DATA_BLOCK "DB823_Error_Metering"   // DB823
TITLE = Faults general at plant and machine
{ S7_Optimized_Access := 'FALSE' }
VERSION : 0.1
   VAR
      FeedPump : Array[0..12] of "UDT1801_FLT_auxDrive";
      EdgeFilter : Array[0..12] of "UDT1801_EdgeFilter";
      MeteringPump : Array[0..12] of "UDT1853_FLT_MeteringPump";   // Metering pump
      Flow_Component : Array[0..12] of "UDT1822_FLT_PV_Flow";   // Process value flow component, mixing ratio
      Pressure_Component : Array[0..12] of "UDT1820_FLT_ProcessValue";   // Process value pressure at metering unit of component
      PrePressure_Component : Array[0..12] of "UDT1820_FLT_ProcessValue";   // Process value pressure at metering unit of component
      MicroMeteringUnit : Array[0..12] of "UDT1807_FaultMicroMeter";   // Micro metering unit ( Color)
      Temperature_HeatexchangerLP : Array[0..12] of "UDT1820_FLT_ProcessValue";   // Process value tempering heat exchanger
      Temperature_HeatexchangerHP : Array[0..12] of "UDT1820_FLT_ProcessValue";   // Process value tempering heat exchanger
      Temperature_Pump : Array[0..12] of "UDT1820_FLT_ProcessValue";   // Process value tempering pumps
      DifferencePressure : Array[0..12] of Struct
         BeforeEdge : "UDT1820_FLT_ProcessValue";
         BehindEdge : "UDT1820_FLT_ProcessValue";
         DifferenceEdge : "UDT1820_FLT_ProcessValue";
         BeforeHP : "UDT1820_FLT_ProcessValue";
         BehindHP : "UDT1820_FLT_ProcessValue";
         DifferenceHP : "UDT1820_FLT_ProcessValue";
      END_STRUCT;
      Heating : Array[0..12] of Struct
         Heating : Array[1..8] of "UDT1804_FLT_Controller";
      END_STRUCT;
   END_VAR
BEGIN
   FeedPump[0].FLT_Motorprotection := FALSE;
   FeedPump[0].FLT_FrequencyConverter := FALSE;
   FeedPump[0].FLT_MaxP_MaxLTripTray := FALSE;
   FeedPump[0].FLT_Dryrunsafety := FALSE;
   FeedPump[0].FLT_wrong_Timevalue := FALSE;
   FeedPump[0].FLT_MaxPressureDiff := FALSE;
   FeedPump[0].Mes_Min_temp := FALSE;
   FeedPump[0].FLT_MotorFan := FALSE;
   FeedPump[0].Mes_Min_Level := FALSE;
   FeedPump[0].FLT_No_Barrel := FALSE;
   FeedPump[0].Mes_No_Barrel := FALSE;
   FeedPump[0].Spare_1_3 := FALSE;
   FeedPump[0].Spare_1_4 := FALSE;
   FeedPump[0].Spare_1_5 := FALSE;
   FeedPump[0].Spare_1_6 := FALSE;
   FeedPump[0].Spare_1_7 := FALSE;
   FeedPump[1].FLT_Motorprotection := FALSE;
   FeedPump[1].FLT_FrequencyConverter := FALSE;
   FeedPump[1].FLT_MaxP_MaxLTripTray := FALSE;
   FeedPump[1].FLT_Dryrunsafety := FALSE;
   FeedPump[1].FLT_wrong_Timevalue := FALSE;
   FeedPump[1].FLT_MaxPressureDiff := FALSE;
   FeedPump[1].Mes_Min_temp := FALSE;
   FeedPump[1].FLT_MotorFan := FALSE;
   FeedPump[1].Mes_Min_Level := FALSE;
   FeedPump[1].FLT_No_Barrel := FALSE;
   FeedPump[1].Mes_No_Barrel := FALSE;
   FeedPump[1].Spare_1_3 := FALSE;
   FeedPump[1].Spare_1_4 := FALSE;
   FeedPump[1].Spare_1_5 := FALSE;
   FeedPump[1].Spare_1_6 := FALSE;
   FeedPump[1].Spare_1_7 := FALSE;
   FeedPump[2].FLT_Motorprotection := FALSE;
   FeedPump[2].FLT_FrequencyConverter := FALSE;
   FeedPump[2].FLT_MaxP_MaxLTripTray := FALSE;
   FeedPump[2].FLT_Dryrunsafety := FALSE;
   FeedPump[2].FLT_wrong_Timevalue := FALSE;
   FeedPump[2].FLT_MaxPressureDiff := FALSE;
   FeedPump[2].Mes_Min_temp := FALSE;
   FeedPump[2].FLT_MotorFan := FALSE;
   FeedPump[2].Mes_Min_Level := FALSE;
   FeedPump[2].FLT_No_Barrel := FALSE;
   FeedPump[2].Mes_No_Barrel := FALSE;
   FeedPump[2].Spare_1_3 := FALSE;
   FeedPump[2].Spare_1_4 := FALSE;
   FeedPump[2].Spare_1_5 := FALSE;
   FeedPump[2].Spare_1_6 := FALSE;
   FeedPump[2].Spare_1_7 := FALSE;
   FeedPump[3].FLT_Motorprotection := FALSE;
   FeedPump[3].FLT_FrequencyConverter := FALSE;
   FeedPump[3].FLT_MaxP_MaxLTripTray := FALSE;
   FeedPump[3].FLT_Dryrunsafety := FALSE;
   FeedPump[3].FLT_wrong_Timevalue := FALSE;
   FeedPump[3].FLT_MaxPressureDiff := FALSE;
   FeedPump[3].Mes_Min_temp := FALSE;
   FeedPump[3].FLT_MotorFan := FALSE;
   FeedPump[3].Mes_Min_Level := FALSE;
   FeedPump[3].FLT_No_Barrel := FALSE;
   FeedPump[3].Mes_No_Barrel := FALSE;
   FeedPump[3].Spare_1_3 := FALSE;
   FeedPump[3].Spare_1_4 := FALSE;
   FeedPump[3].Spare_1_5 := FALSE;
   FeedPump[3].Spare_1_6 := FALSE;
   FeedPump[3].Spare_1_7 := FALSE;
   FeedPump[4].FLT_Motorprotection := FALSE;
   FeedPump[4].FLT_FrequencyConverter := FALSE;
   FeedPump[4].FLT_MaxP_MaxLTripTray := FALSE;
   FeedPump[4].FLT_Dryrunsafety := FALSE;
   FeedPump[4].FLT_wrong_Timevalue := FALSE;
   FeedPump[4].FLT_MaxPressureDiff := FALSE;
   FeedPump[4].Mes_Min_temp := FALSE;
   FeedPump[4].FLT_MotorFan := FALSE;
   FeedPump[4].Mes_Min_Level := FALSE;
   FeedPump[4].FLT_No_Barrel := FALSE;
   FeedPump[4].Mes_No_Barrel := FALSE;
   FeedPump[4].Spare_1_3 := FALSE;
   FeedPump[4].Spare_1_4 := FALSE;
   FeedPump[4].Spare_1_5 := FALSE;
   FeedPump[4].Spare_1_6 := FALSE;
   FeedPump[4].Spare_1_7 := FALSE;
   FeedPump[5].FLT_Motorprotection := FALSE;
   FeedPump[5].FLT_FrequencyConverter := FALSE;
   FeedPump[5].FLT_MaxP_MaxLTripTray := FALSE;
   FeedPump[5].FLT_Dryrunsafety := FALSE;
   FeedPump[5].FLT_wrong_Timevalue := FALSE;
   FeedPump[5].FLT_MaxPressureDiff := FALSE;
   FeedPump[5].Mes_Min_temp := FALSE;
   FeedPump[5].FLT_MotorFan := FALSE;
   FeedPump[5].Mes_Min_Level := FALSE;
   FeedPump[5].FLT_No_Barrel := FALSE;
   FeedPump[5].Mes_No_Barrel := FALSE;
   FeedPump[5].Spare_1_3 := FALSE;
   FeedPump[5].Spare_1_4 := FALSE;
   FeedPump[5].Spare_1_5 := FALSE;
   FeedPump[5].Spare_1_6 := FALSE;
   FeedPump[5].Spare_1_7 := FALSE;
   FeedPump[6].FLT_Motorprotection := FALSE;
   FeedPump[6].FLT_FrequencyConverter := FALSE;
   FeedPump[6].FLT_MaxP_MaxLTripTray := FALSE;
   FeedPump[6].FLT_Dryrunsafety := FALSE;
   FeedPump[6].FLT_wrong_Timevalue := FALSE;
   FeedPump[6].FLT_MaxPressureDiff := FALSE;
   FeedPump[6].Mes_Min_temp := FALSE;
   FeedPump[6].FLT_MotorFan := FALSE;
   FeedPump[6].Mes_Min_Level := FALSE;
   FeedPump[6].FLT_No_Barrel := FALSE;
   FeedPump[6].Mes_No_Barrel := FALSE;
   FeedPump[6].Spare_1_3 := FALSE;
   FeedPump[6].Spare_1_4 := FALSE;
   FeedPump[6].Spare_1_5 := FALSE;
   FeedPump[6].Spare_1_6 := FALSE;
   FeedPump[6].Spare_1_7 := FALSE;
   FeedPump[7].FLT_Motorprotection := FALSE;
   FeedPump[7].FLT_FrequencyConverter := FALSE;
   FeedPump[7].FLT_MaxP_MaxLTripTray := FALSE;
   FeedPump[7].FLT_Dryrunsafety := FALSE;
   FeedPump[7].FLT_wrong_Timevalue := FALSE;
   FeedPump[7].FLT_MaxPressureDiff := FALSE;
   FeedPump[7].Mes_Min_temp := FALSE;
   FeedPump[7].FLT_MotorFan := FALSE;
   FeedPump[7].Mes_Min_Level := FALSE;
   FeedPump[7].FLT_No_Barrel := FALSE;
   FeedPump[7].Mes_No_Barrel := FALSE;
   FeedPump[7].Spare_1_3 := FALSE;
   FeedPump[7].Spare_1_4 := FALSE;
   FeedPump[7].Spare_1_5 := FALSE;
   FeedPump[7].Spare_1_6 := FALSE;
   FeedPump[7].Spare_1_7 := FALSE;
   FeedPump[8].FLT_Motorprotection := FALSE;
   FeedPump[8].FLT_FrequencyConverter := FALSE;
   FeedPump[8].FLT_MaxP_MaxLTripTray := FALSE;
   FeedPump[8].FLT_Dryrunsafety := FALSE;
   FeedPump[8].FLT_wrong_Timevalue := FALSE;
   FeedPump[8].FLT_MaxPressureDiff := FALSE;
   FeedPump[8].Mes_Min_temp := FALSE;
   FeedPump[8].FLT_MotorFan := FALSE;
   FeedPump[8].Mes_Min_Level := FALSE;
   FeedPump[8].FLT_No_Barrel := FALSE;
   FeedPump[8].Mes_No_Barrel := FALSE;
   FeedPump[8].Spare_1_3 := FALSE;
   FeedPump[8].Spare_1_4 := FALSE;
   FeedPump[8].Spare_1_5 := FALSE;
   FeedPump[8].Spare_1_6 := FALSE;
   FeedPump[8].Spare_1_7 := FALSE;
   FeedPump[9].FLT_Motorprotection := FALSE;
   FeedPump[9].FLT_FrequencyConverter := FALSE;
   FeedPump[9].FLT_MaxP_MaxLTripTray := FALSE;
   FeedPump[9].FLT_Dryrunsafety := FALSE;
   FeedPump[9].FLT_wrong_Timevalue := FALSE;
   FeedPump[9].FLT_MaxPressureDiff := FALSE;
   FeedPump[9].Mes_Min_temp := FALSE;
   FeedPump[9].FLT_MotorFan := FALSE;
   FeedPump[9].Mes_Min_Level := FALSE;
   FeedPump[9].FLT_No_Barrel := FALSE;
   FeedPump[9].Mes_No_Barrel := FALSE;
   FeedPump[9].Spare_1_3 := FALSE;
   FeedPump[9].Spare_1_4 := FALSE;
   FeedPump[9].Spare_1_5 := FALSE;
   FeedPump[9].Spare_1_6 := FALSE;
   FeedPump[9].Spare_1_7 := FALSE;
   FeedPump[10].FLT_Motorprotection := FALSE;
   FeedPump[10].FLT_FrequencyConverter := FALSE;
   FeedPump[10].FLT_MaxP_MaxLTripTray := FALSE;
   FeedPump[10].FLT_Dryrunsafety := FALSE;
   FeedPump[10].FLT_wrong_Timevalue := FALSE;
   FeedPump[10].FLT_MaxPressureDiff := FALSE;
   FeedPump[10].Mes_Min_temp := FALSE;
   FeedPump[10].FLT_MotorFan := FALSE;
   FeedPump[10].Mes_Min_Level := FALSE;
   FeedPump[10].FLT_No_Barrel := FALSE;
   FeedPump[10].Mes_No_Barrel := FALSE;
   FeedPump[10].Spare_1_3 := FALSE;
   FeedPump[10].Spare_1_4 := FALSE;
   FeedPump[10].Spare_1_5 := FALSE;
   FeedPump[10].Spare_1_6 := FALSE;
   FeedPump[10].Spare_1_7 := FALSE;
   FeedPump[11].FLT_Motorprotection := FALSE;
   FeedPump[11].FLT_FrequencyConverter := FALSE;
   FeedPump[11].FLT_MaxP_MaxLTripTray := FALSE;
   FeedPump[11].FLT_Dryrunsafety := FALSE;
   FeedPump[11].FLT_wrong_Timevalue := FALSE;
   FeedPump[11].FLT_MaxPressureDiff := FALSE;
   FeedPump[11].Mes_Min_temp := FALSE;
   FeedPump[11].FLT_MotorFan := FALSE;
   FeedPump[11].Mes_Min_Level := FALSE;
   FeedPump[11].FLT_No_Barrel := FALSE;
   FeedPump[11].Mes_No_Barrel := FALSE;
   FeedPump[11].Spare_1_3 := FALSE;
   FeedPump[11].Spare_1_4 := FALSE;
   FeedPump[11].Spare_1_5 := FALSE;
   FeedPump[11].Spare_1_6 := FALSE;
   FeedPump[11].Spare_1_7 := FALSE;
   FeedPump[12].FLT_Motorprotection := FALSE;
   FeedPump[12].FLT_FrequencyConverter := FALSE;
   FeedPump[12].FLT_MaxP_MaxLTripTray := FALSE;
   FeedPump[12].FLT_Dryrunsafety := FALSE;
   FeedPump[12].FLT_wrong_Timevalue := FALSE;
   FeedPump[12].FLT_MaxPressureDiff := FALSE;
   FeedPump[12].Mes_Min_temp := FALSE;
   FeedPump[12].FLT_MotorFan := FALSE;
   // 3232 more start values not shown
END_DATA_BLOCK

DATA_BLOCK "DB824_Error_MH_CP"   // DB824
TITLE = Faults mixinghead and cleaning piston
{ S7_Optimized_Access := 'FALSE' }
VERSION : 0.1
   VAR
      MH_Control : Array[0..16] of "UDT1842_FLT_MH_Control";
      CPiston : Array[0..16] of "UDT1871_FLT_CPiston";
      Temperature : Array[1..6, 0..16] of "UDT1820_FLT_ProcessValue";
      Pressure : Array[1..6, 0..16] of "UDT1820_FLT_ProcessValue";
      SteeringPiston : Array[0..16] of "UDT1820_FLT_ProcessValue";
      CleaningPiston : Array[0..16] of "UDT1820_FLT_ProcessValue";
      InertingBlowOut_MH : Array[0..16] of "UDT1825_FLT_Inerting";
      EmergencyStop_Opanel_MH : Array[1..32] of Bool;
   END_VAR
BEGIN
   MH_Control[0].FLT_MH_dontOpen := FALSE;
   MH_Control[0].FLT_MH_dontClose := FALSE;
   MH_Control[0].FLT_ShotStopped := FALSE;
   MH_Control[0].FLT_MH_OpenWOactivation := FALSE;
   MH_Control[0].FLT_MH_CloseDuringShot := FALSE;
   MH_Control[0].WRN_ShotTimeShort := FALSE;
   MH_Control[0].WRN_ShotTimeLong := FALSE;
   MH_Control[0].FLT_ShotTimeShort := FALSE;
   MH_Control[0].FLT_MH_bounce := FALSE;
   MH_Control[0].FLT_RT_Lock := FALSE;
   MH_Control[0].FLT_RT_Unlock := FALSE;
   MH_Control[0].WRN_NozzleLeakageTest_active := FALSE;
   MH_Control[0].Spare_1_4 := FALSE;
   MH_Control[0].Spare_1_5 := FALSE;
   MH_Control[0].Spare_1_6 := FALSE;
   MH_Control[0].FLTCompNotOnThisMH := FALSE;
   MH_Control[1].FLT_MH_dontOpen := FALSE;
   MH_Control[1].FLT_MH_dontClose := FALSE;
   MH_Control[1].FLT_ShotStopped := FALSE;
   MH_Control[1].FLT_MH_OpenWOactivation := FALSE;
   MH_Control[1].FLT_MH_CloseDuringShot := FALSE;
   MH_Control[1].WRN_ShotTimeShort := FALSE;
   MH_Control[1].WRN_ShotTimeLong := FALSE;
   MH_Control[1].FLT_ShotTimeShort := FALSE;
   MH_Control[1].FLT_MH_bounce := FALSE;
   MH_Control[1].FLT_RT_Lock := FALSE;
   MH_Control[1].FLT_RT_Unlock := FALSE;
   MH_Control[1].WRN_NozzleLeakageTest_active := FALSE;
   MH_Control[1].Spare_1_4 := FALSE;
   MH_Control[1].Spare_1_5 := FALSE;
   MH_Control[1].Spare_1_6 := FALSE;
   MH_Control[1].FLTCompNotOnThisMH := FALSE;
   MH_Control[2].FLT_MH_dontOpen := FALSE;
   MH_Control[2].FLT_MH_dontClose := FALSE;
   MH_Control[2].FLT_ShotStopped := FALSE;
   MH_Control[2].FLT_MH_OpenWOactivation := FALSE;
   MH_Control[2].FLT_MH_CloseDuringShot := FALSE;
   MH_Control[2].WRN_ShotTimeShort := FALSE;
   MH_Control[2].WRN_ShotTimeLong := FALSE;
   MH_Control[2].FLT_ShotTimeShort := FALSE;
   MH_Control[2].FLT_MH_bounce := FALSE;
   MH_Control[2].FLT_RT_Lock := FALSE;
   MH_Control[2].FLT_RT_Unlock := FALSE;
   MH_Control[2].WRN_NozzleLeakageTest_active := FALSE;
   MH_Control[2].Spare_1_4 := FALSE;
   MH_Control[2].Spare_1_5 := FALSE;
   MH_Control[2].Spare_1_6 := FALSE;
   MH_Control[2].FLTCompNotOnThisMH := FALSE;
   MH_Control[3].FLT_MH_dontOpen := FALSE;
   MH_Control[3].FLT_MH_dontClose := FALSE;
   MH_Control[3].FLT_ShotStopped := FALSE;
   MH_Control[3].FLT_MH_OpenWOactivation := FALSE;
   MH_Control[3].FLT_MH_CloseDuringShot := FALSE;
   MH_Control[3].WRN_ShotTimeShort := FALSE;
   MH_Control[3].WRN_ShotTimeLong := FALSE;
   MH_Control[3].FLT_ShotTimeShort := FALSE;
   MH_Control[3].FLT_MH_bounce := FALSE;
   MH_Control[3].FLT_RT_Lock := FALSE;
   MH_Control[3].FLT_RT_Unlock := FALSE;
   MH_Control[3].WRN_NozzleLeakageTest_active := FALSE;
   MH_Control[3].Spare_1_4 := FALSE;
   MH_Control[3].Spare_1_5 := FALSE;
   MH_Control[3].Spare_1_6 := FALSE;
   MH_Control[3].FLTCompNotOnThisMH := FALSE;
   MH_Control[4].FLT_MH_dontOpen := FALSE;
   MH_Control[4].FLT_MH_dontClose := FALSE;
   MH_Control[4].FLT_ShotStopped := FALSE;
   MH_Control[4].FLT_MH_OpenWOactivation := FALSE;
   MH_Control[4].FLT_MH_CloseDuringShot := FALSE;
   MH_Control[4].WRN_ShotTimeShort := FALSE;
   MH_Control[4].WRN_ShotTimeLong := FALSE;
   MH_Control[4].FLT_ShotTimeShort := FALSE;
   MH_Control[4].FLT_MH_bounce := FALSE;
   MH_Control[4].FLT_RT_Lock := FALSE;
   MH_Control[4].FLT_RT_Unlock := FALSE;
   MH_Control[4].WRN_NozzleLeakageTest_active := FALSE;
   MH_Control[4].Spare_1_4 := FALSE;
   MH_Control[4].Spare_1_5 := FALSE;
   MH_Control[4].Spare_1_6 := FALSE;
   MH_Control[4].FLTCompNotOnThisMH := FALSE;
   MH_Control[5].FLT_MH_dontOpen := FALSE;
   MH_Control[5].FLT_MH_dontClose := FALSE;
   MH_Control[5].FLT_ShotStopped := FALSE;
   MH_Control[5].FLT_MH_OpenWOactivation := FALSE;
   MH_Control[5].FLT_MH_CloseDuringShot := FALSE;
   MH_Control[5].WRN_ShotTimeShort := FALSE;
   MH_Control[5].WRN_ShotTimeLong := FALSE;
   MH_Control[5].FLT_ShotTimeShort := FALSE;
   MH_Control[5].FLT_MH_bounce := FALSE;
   MH_Control[5].FLT_RT_Lock := FALSE;
   MH_Control[5].FLT_RT_Unlock := FALSE;
   MH_Control[5].WRN_NozzleLeakageTest_active := FALSE;
   MH_Control[5].Spare_1_4 := FALSE;
   MH_Control[5].Spare_1_5 := FALSE;
   MH_Control[5].Spare_1_6 := FALSE;
   MH_Control[5].FLTCompNotOnThisMH := FALSE;
   MH_Control[6].FLT_MH_dontOpen := FALSE;
   MH_Control[6].FLT_MH_dontClose := FALSE;
   MH_Control[6].FLT_ShotStopped := FALSE;
   MH_Control[6].FLT_MH_OpenWOactivation := FALSE;
   MH_Control[6].FLT_MH_CloseDuringShot := FALSE;
   MH_Control[6].WRN_ShotTimeShort := FALSE;
   MH_Control[6].WRN_ShotTimeLong := FALSE;
   MH_Control[6].FLT_ShotTimeShort := FALSE;
   MH_Control[6].FLT_MH_bounce := FALSE;
   MH_Control[6].FLT_RT_Lock := FALSE;
   MH_Control[6].FLT_RT_Unlock := FALSE;
   MH_Control[6].WRN_NozzleLeakageTest_active := FALSE;
   MH_Control[6].Spare_1_4 := FALSE;
   MH_Control[6].Spare_1_5 := FALSE;
   MH_Control[6].Spare_1_6 := FALSE;
   MH_Control[6].FLTCompNotOnThisMH := FALSE;
   MH_Control[7].FLT_MH_dontOpen := FALSE;
   MH_Control[7].FLT_MH_dontClose := FALSE;
   MH_Control[7].FLT_ShotStopped := FALSE;
   MH_Control[7].FLT_MH_OpenWOactivation := FALSE;
   MH_Control[7].FLT_MH_CloseDuringShot := FALSE;
   MH_Control[7].WRN_ShotTimeShort := FALSE;
   MH_Control[7].WRN_ShotTimeLong := FALSE;
   MH_Control[7].FLT_ShotTimeShort := FALSE;
   MH_Control[7].FLT_MH_bounce := FALSE;
   MH_Control[7].FLT_RT_Lock := FALSE;
   MH_Control[7].FLT_RT_Unlock := FALSE;
   MH_Control[7].WRN_NozzleLeakageTest_active := FALSE;
   MH_Control[7].Spare_1_4 := FALSE;
   MH_Control[7].Spare_1_5 := FALSE;
   MH_Control[7].Spare_1_6 := FALSE;
   MH_Control[7].FLTCompNotOnThisMH := FALSE;
   MH_Control[8].FLT_MH_dontOpen := FALSE;
   MH_Control[8].FLT_MH_dontClose := FALSE;
   MH_Control[8].FLT_ShotStopped := FALSE;
   MH_Control[8].FLT_MH_OpenWOactivation := FALSE;
   MH_Control[8].FLT_MH_CloseDuringShot := FALSE;
   MH_Control[8].WRN_ShotTimeShort := FALSE;
   MH_Control[8].WRN_ShotTimeLong := FALSE;
   MH_Control[8].FLT_ShotTimeShort := FALSE;
   MH_Control[8].FLT_MH_bounce := FALSE;
   MH_Control[8].FLT_RT_Lock := FALSE;
   MH_Control[8].FLT_RT_Unlock := FALSE;
   MH_Control[8].WRN_NozzleLeakageTest_active := FALSE;
   MH_Control[8].Spare_1_4 := FALSE;
   MH_Control[8].Spare_1_5 := FALSE;
   MH_Control[8].Spare_1_6 := FALSE;
   MH_Control[8].FLTCompNotOnThisMH := FALSE;
   MH_Control[9].FLT_MH_dontOpen := FALSE;
   MH_Control[9].FLT_MH_dontClose := FALSE;
   MH_Control[9].FLT_ShotStopped := FALSE;
   MH_Control[9].FLT_MH_OpenWOactivation := FALSE;
   MH_Control[9].FLT_MH_CloseDuringShot := FALSE;
   MH_Control[9].WRN_ShotTimeShort := FALSE;
   MH_Control[9].WRN_ShotTimeLong := FALSE;
   MH_Control[9].FLT_ShotTimeShort := FALSE;
   MH_Control[9].FLT_MH_bounce := FALSE;
   MH_Control[9].FLT_RT_Lock := FALSE;
   MH_Control[9].FLT_RT_Unlock := FALSE;
   MH_Control[9].WRN_NozzleLeakageTest_active := FALSE;
   MH_Control[9].Spare_1_4 := FALSE;
   MH_Control[9].Spare_1_5 := FALSE;
   MH_Control[9].Spare_1_6 := FALSE;
   MH_Control[9].FLTCompNotOnThisMH := FALSE;
   MH_Control[10].FLT_MH_dontOpen := FALSE;
   MH_Control[10].FLT_MH_dontClose := FALSE;
   MH_Control[10].FLT_ShotStopped := FALSE;
   MH_Control[10].FLT_MH_OpenWOactivation := FALSE;
   MH_Control[10].FLT_MH_CloseDuringShot := FALSE;
   MH_Control[10].WRN_ShotTimeShort := FALSE;
   MH_Control[10].WRN_ShotTimeLong := FALSE;
   MH_Control[10].FLT_ShotTimeShort := FALSE;
   MH_Control[10].FLT_MH_bounce := FALSE;
   MH_Control[10].FLT_RT_Lock := FALSE;
   MH_Control[10].FLT_RT_Unlock := FALSE;
   MH_Control[10].WRN_NozzleLeakageTest_active := FALSE;
   MH_Control[10].Spare_1_4 := FALSE;
   MH_Control[10].Spare_1_5 := FALSE;
   MH_Control[10].Spare_1_6 := FALSE;
   MH_Control[10].FLTCompNotOnThisMH := FALSE;
   MH_Control[11].FLT_MH_dontOpen := FALSE;
   MH_Control[11].FLT_MH_dontClose := FALSE;
   MH_Control[11].FLT_ShotStopped := FALSE;
   MH_Control[11].FLT_MH_OpenWOactivation := FALSE;
   MH_Control[11].FLT_MH_CloseDuringShot := FALSE;
   MH_Control[11].WRN_ShotTimeShort := FALSE;
   MH_Control[11].WRN_ShotTimeLong := FALSE;
   MH_Control[11].FLT_ShotTimeShort := FALSE;
   MH_Control[11].FLT_MH_bounce := FALSE;
   MH_Control[11].FLT_RT_Lock := FALSE;
   MH_Control[11].FLT_RT_Unlock := FALSE;
   MH_Control[11].WRN_NozzleLeakageTest_active := FALSE;
   MH_Control[11].Spare_1_4 := FALSE;
   MH_Control[11].Spare_1_5 := FALSE;
   MH_Control[11].Spare_1_6 := FALSE;
   MH_Control[11].FLTCompNotOnThisMH := FALSE;
   MH_Control[12].FLT_MH_dontOpen := FALSE;
   MH_Control[12].FLT_MH_dontClose := FALSE;
   MH_Control[12].FLT_ShotStopped := FALSE;
   MH_Control[12].FLT_MH_OpenWOactivation := FALSE;
   MH_Control[12].FLT_MH_CloseDuringShot := FALSE;
   MH_Control[12].WRN_ShotTimeShort := FALSE;
   MH_Control[12].WRN_ShotTimeLong := FALSE;
   MH_Control[12].FLT_ShotTimeShort := FALSE;
   // 4320 more start values not shown
END_DATA_BLOCK

DATA_BLOCK "DB825_Error_Interface"   // DB825
TITLE = Faults general at plant and machine
{ S7_Optimized_Access := 'FALSE' }
VERSION : 0.1
   VAR
      Interface_MC : Array[1..16] of "UDT1816_FLT_IF_SP_MC";   // Interface between pouring machine and mould carrier
      Interface_externalPlant : Array[1..16] of "UDT1817_FLT_IF_extPlant";   // Interface between pouring machine and external plant
      EmergencyStop_MC : Array[1..16] of Bool;   // Emergency stop button actuated
   END_VAR
BEGIN
   Interface_MC[1].Fault_IF := FALSE;
   Interface_MC[1].FLT_pouring_release := FALSE;
   Interface_MC[1].FLT_SWU_release := FALSE;
   Interface_MC[1].FLT_Stop_while_selected := FALSE;
   Interface_MC[1].FLT_op_mode_O := FALSE;
   Interface_MC[1].FLT_Cycle_release := FALSE;
   Interface_MC[1].FLT_Communication := FALSE;
   Interface_MC[1].FLT_NoCupAtTestshotposition := FALSE;
   Interface_MC[1].Spare_1_0 := FALSE;
   Interface_MC[1].Spare_1_1 := FALSE;
   Interface_MC[1].Spare_1_2 := FALSE;
   Interface_MC[1].Spare_1_3 := FALSE;
   Interface_MC[1].Spare_1_4 := FALSE;
   Interface_MC[1].Spare_1_5 := FALSE;
   Interface_MC[1].Spare_1_6 := FALSE;
   Interface_MC[1].Spare_1_7 := FALSE;
   Interface_MC[2].Fault_IF := FALSE;
   Interface_MC[2].FLT_pouring_release := FALSE;
   Interface_MC[2].FLT_SWU_release := FALSE;
   Interface_MC[2].FLT_Stop_while_selected := FALSE;
   Interface_MC[2].FLT_op_mode_O := FALSE;
   Interface_MC[2].FLT_Cycle_release := FALSE;
   Interface_MC[2].FLT_Communication := FALSE;
   Interface_MC[2].FLT_NoCupAtTestshotposition := FALSE;
   Interface_MC[2].Spare_1_0 := FALSE;
   Interface_MC[2].Spare_1_1 := FALSE;
   Interface_MC[2].Spare_1_2 := FALSE;
   Interface_MC[2].Spare_1_3 := FALSE;
   Interface_MC[2].Spare_1_4 := FALSE;
   Interface_MC[2].Spare_1_5 := FALSE;
   Interface_MC[2].Spare_1_6 := FALSE;
   Interface_MC[2].Spare_1_7 := FALSE;
   Interface_MC[3].Fault_IF := FALSE;
   Interface_MC[3].FLT_pouring_release := FALSE;
   Interface_MC[3].FLT_SWU_release := FALSE;
   Interface_MC[3].FLT_Stop_while_selected := FALSE;
   Interface_MC[3].FLT_op_mode_O := FALSE;
   Interface_MC[3].FLT_Cycle_release := FALSE;
   Interface_MC[3].FLT_Communication := FALSE;
   Interface_MC[3].FLT_NoCupAtTestshotposition := FALSE;
   Interface_MC[3].Spare_1_0 := FALSE;
   Interface_MC[3].Spare_1_1 := FALSE;
   Interface_MC[3].Spare_1_2 := FALSE;
   Interface_MC[3].Spare_1_3 := FALSE;
   Interface_MC[3].Spare_1_4 := FALSE;
   Interface_MC[3].Spare_1_5 := FALSE;
   Interface_MC[3].Spare_1_6 := FALSE;
   Interface_MC[3].Spare_1_7 := FALSE;
   Interface_MC[4].Fault_IF := FALSE;
   Interface_MC[4].FLT_pouring_release := FALSE;
   Interface_MC[4].FLT_SWU_release := FALSE;
   Interface_MC[4].FLT_Stop_while_selected := FALSE;
   Interface_MC[4].FLT_op_mode_O := FALSE;
   Interface_MC[4].FLT_Cycle_release := FALSE;
   Interface_MC[4].FLT_Communication := FALSE;
   Interface_MC[4].FLT_NoCupAtTestshotposition := FALSE;
   Interface_MC[4].Spare_1_0 := FALSE;
   Interface_MC[4].Spare_1_1 := FALSE;
   Interface_MC[4].Spare_1_2 := FALSE;
   Interface_MC[4].Spare_1_3 := FALSE;
   Interface_MC[4].Spare_1_4 := FALSE;
   Interface_MC[4].Spare_1_5 := FALSE;
   Interface_MC[4].Spare_1_6 := FALSE;
   Interface_MC[4].Spare_1_7 := FALSE;
   Interface_MC[5].Fault_IF := FALSE;
   Interface_MC[5].FLT_pouring_release := FALSE;
   Interface_MC[5].FLT_SWU_release := FALSE;
   Interface_MC[5].FLT_Stop_while_selected := FALSE;
   Interface_MC[5].FLT_op_mode_O := FALSE;
   Interface_MC[5].FLT_Cycle_release := FALSE;
   Interface_MC[5].FLT_Communication := FALSE;
   Interface_MC[5].FLT_NoCupAtTestshotposition := FALSE;
   Interface_MC[5].Spare_1_0 := FALSE;
   Interface_MC[5].Spare_1_1 := FALSE;
   Interface_MC[5].Spare_1_2 := FALSE;
   Interface_MC[5].Spare_1_3 := FALSE;
   Interface_MC[5].Spare_1_4 := FALSE;
   Interface_MC[5].Spare_1_5 := FALSE;
   Interface_MC[5].Spare_1_6 := FALSE;
   Interface_MC[5].Spare_1_7 := FALSE;
   Interface_MC[6].Fault_IF := FALSE;
   Interface_MC[6].FLT_pouring_release := FALSE;
   Interface_MC[6].FLT_SWU_release := FALSE;
   Interface_MC[6].FLT_Stop_while_selected := FALSE;
   Interface_MC[6].FLT_op_mode_O := FALSE;
   Interface_MC[6].FLT_Cycle_release := FALSE;
   Interface_MC[6].FLT_Communication := FALSE;
   Interface_MC[6].FLT_NoCupAtTestshotposition := FALSE;
   Interface_MC[6].Spare_1_0 := FALSE;
   Interface_MC[6].Spare_1_1 := FALSE;
   Interface_MC[6].Spare_1_2 := FALSE;
   Interface_MC[6].Spare_1_3 := FALSE;
   Interface_MC[6].Spare_1_4 := FALSE;
   Interface_MC[6].Spare_1_5 := FALSE;
   Interface_MC[6].Spare_1_6 := FALSE;
   Interface_MC[6].Spare_1_7 := FALSE;
   Interface_MC[7].Fault_IF := FALSE;
   Interface_MC[7].FLT_pouring_release := FALSE;
   Interface_MC[7].FLT_SWU_release := FALSE;
   Interface_MC[7].FLT_Stop_while_selected := FALSE;
   Interface_MC[7].FLT_op_mode_O := FALSE;
   Interface_MC[7].FLT_Cycle_release := FALSE;
   Interface_MC[7].FLT_Communication := FALSE;
   Interface_MC[7].FLT_NoCupAtTestshotposition := FALSE;
   Interface_MC[7].Spare_1_0 := FALSE;
   Interface_MC[7].Spare_1_1 := FALSE;
   Interface_MC[7].Spare_1_2 := FALSE;
   Interface_MC[7].Spare_1_3 := FALSE;
   Interface_MC[7].Spare_1_4 := FALSE;
   Interface_MC[7].Spare_1_5 := FALSE;
   Interface_MC[7].Spare_1_6 := FALSE;
   Interface_MC[7].Spare_1_7 := FALSE;
   Interface_MC[8].Fault_IF := FALSE;
   Interface_MC[8].FLT_pouring_release := FALSE;
   Interface_MC[8].FLT_SWU_release := FALSE;
   Interface_MC[8].FLT_Stop_while_selected := FALSE;
   Interface_MC[8].FLT_op_mode_O := FALSE;
   Interface_MC[8].FLT_Cycle_release := FALSE;
   Interface_MC[8].FLT_Communication := FALSE;
   Interface_MC[8].FLT_NoCupAtTestshotposition := FALSE;
   Interface_MC[8].Spare_1_0 := FALSE;
   Interface_MC[8].Spare_1_1 := FALSE;
   Interface_MC[8].Spare_1_2 := FALSE;
   Interface_MC[8].Spare_1_3 := FALSE;
   Interface_MC[8].Spare_1_4 := FALSE;
   Interface_MC[8].Spare_1_5 := FALSE;
   Interface_MC[8].Spare_1_6 := FALSE;
   Interface_MC[8].Spare_1_7 := FALSE;
   Interface_MC[9].Fault_IF := FALSE;
   Interface_MC[9].FLT_pouring_release := FALSE;
   Interface_MC[9].FLT_SWU_release := FALSE;
   Interface_MC[9].FLT_Stop_while_selected := FALSE;
   Interface_MC[9].FLT_op_mode_O := FALSE;
   Interface_MC[9].FLT_Cycle_release := FALSE;
   Interface_MC[9].FLT_Communication := FALSE;
   Interface_MC[9].FLT_NoCupAtTestshotposition := FALSE;
   Interface_MC[9].Spare_1_0 := FALSE;
   Interface_MC[9].Spare_1_1 := FALSE;
   Interface_MC[9].Spare_1_2 := FALSE;
   Interface_MC[9].Spare_1_3 := FALSE;
   Interface_MC[9].Spare_1_4 := FALSE;
   Interface_MC[9].Spare_1_5 := FALSE;
   Interface_MC[9].Spare_1_6 := FALSE;
   Interface_MC[9].Spare_1_7 := FALSE;
   Interface_MC[10].Fault_IF := FALSE;
   Interface_MC[10].FLT_pouring_release := FALSE;
   Interface_MC[10].FLT_SWU_release := FALSE;
   Interface_MC[10].FLT_Stop_while_selected := FALSE;
   Interface_MC[10].FLT_op_mode_O := FALSE;
   Interface_MC[10].FLT_Cycle_release := FALSE;
   Interface_MC[10].FLT_Communication := FALSE;
   Interface_MC[10].FLT_NoCupAtTestshotposition := FALSE;
   Interface_MC[10].Spare_1_0 := FALSE;
   Interface_MC[10].Spare_1_1 := FALSE;
   Interface_MC[10].Spare_1_2 := FALSE;
   Interface_MC[10].Spare_1_3 := FALSE;
   Interface_MC[10].Spare_1_4 := FALSE;
   Interface_MC[10].Spare_1_5 := FALSE;
   Interface_MC[10].Spare_1_6 := FALSE;
   Interface_MC[10].Spare_1_7 := FALSE;
   Interface_MC[11].Fault_IF := FALSE;
   Interface_MC[11].FLT_pouring_release := FALSE;
   Interface_MC[11].FLT_SWU_release := FALSE;
   Interface_MC[11].FLT_Stop_while_selected := FALSE;
   Interface_MC[11].FLT_op_mode_O := FALSE;
   Interface_MC[11].FLT_Cycle_release := FALSE;
   Interface_MC[11].FLT_Communication := FALSE;
   Interface_MC[11].FLT_NoCupAtTestshotposition := FALSE;
   Interface_MC[11].Spare_1_0 := FALSE;
   Interface_MC[11].Spare_1_1 := FALSE;
   Interface_MC[11].Spare_1_2 := FALSE;
   Interface_MC[11].Spare_1_3 := FALSE;
   Interface_MC[11].Spare_1_4 := FALSE;
   Interface_MC[11].Spare_1_5 := FALSE;
   Interface_MC[11].Spare_1_6 := FALSE;
   Interface_MC[11].Spare_1_7 := FALSE;
   Interface_MC[12].Fault_IF := FALSE;
   Interface_MC[12].FLT_pouring_release := FALSE;
   Interface_MC[12].FLT_SWU_release := FALSE;
   Interface_MC[12].FLT_Stop_while_selected := FALSE;
   Interface_MC[12].FLT_op_mode_O := FALSE;
   Interface_MC[12].FLT_Cycle_release := FALSE;
   Interface_MC[12].FLT_Communication := FALSE;
   Interface_MC[12].FLT_NoCupAtTestshotposition := FALSE;
   Interface_MC[12].Spare_1_0 := FALSE;
   Interface_MC[12].Spare_1_1 := FALSE;
   Interface_MC[12].Spare_1_2 := FALSE;
   Interface_MC[12].Spare_1_3 := FALSE;
   Interface_MC[12].Spare_1_4 := FALSE;
   Interface_MC[12].Spare_1_5 := FALSE;
   Interface_MC[12].Spare_1_6 := FALSE;
   Interface_MC[12].Spare_1_7 := FALSE;
   Interface_MC[13].Fault_IF := FALSE;
   Interface_MC[13].FLT_pouring_release := FALSE;
   Interface_MC[13].FLT_SWU_release := FALSE;
   Interface_MC[13].FLT_Stop_while_selected := FALSE;
   Interface_MC[13].FLT_op_mode_O := FALSE;
   Interface_MC[13].FLT_Cycle_release := FALSE;
   Interface_MC[13].FLT_Communication := FALSE;
   Interface_MC[13].FLT_NoCupAtTestshotposition := FALSE;
   // 328 more start values not shown
END_DATA_BLOCK

DATA_BLOCK "DB829_Error_Machine"   // DB829
TITLE = Faults general at plant and machine
{ S7_Optimized_Access := 'FALSE' }
VERSION : 0.1
   VAR
      SWU : Array[1..2] of "UDT1841_FLT_SWU";   // Switch over unit at machine
      PouringCycle : Array[1..2] of "UDT1819_FLT_PouringCycle";   // Pouring cycle
      Foaming_Time : Array[1..2] of "UDT1820_FLT_ProcessValue";   // Process value foaming time
   END_VAR
BEGIN
   SWU[1].FLT_open_SWU_disabelt := FALSE;
   SWU[1].FLT_No_SWU_selected := FALSE;
   SWU[1].FLT_Sel_SWU_not_released := FALSE;
   SWU[1].spare_0_3 := FALSE;
   SWU[1].spare_0_4 := FALSE;
   SWU[1].spare_0_5 := FALSE;
   SWU[1].spare_0_6 := FALSE;
   SWU[1].spare_0_7 := FALSE;
   SWU[1].spare_1_0 := FALSE;
   SWU[1].spare_1_1 := FALSE;
   SWU[1].spare_1_2 := FALSE;
   SWU[1].spare_1_3 := FALSE;
   SWU[1].spare_1_4 := FALSE;
   SWU[1].spare_1_5 := FALSE;
   SWU[1].spare_1_6 := FALSE;
   SWU[1].spare_1_7 := FALSE;
   SWU[2].FLT_open_SWU_disabelt := FALSE;
   SWU[2].FLT_No_SWU_selected := FALSE;
   SWU[2].FLT_Sel_SWU_not_released := FALSE;
   SWU[2].spare_0_3 := FALSE;
   SWU[2].spare_0_4 := FALSE;
   SWU[2].spare_0_5 := FALSE;
   SWU[2].spare_0_6 := FALSE;
   SWU[2].spare_0_7 := FALSE;
   SWU[2].spare_1_0 := FALSE;
   SWU[2].spare_1_1 := FALSE;
   SWU[2].spare_1_2 := FALSE;
   SWU[2].spare_1_3 := FALSE;
   SWU[2].spare_1_4 := FALSE;
   SWU[2].spare_1_5 := FALSE;
   SWU[2].spare_1_6 := FALSE;
   SWU[2].spare_1_7 := FALSE;
   PouringCycle[1].FLT_KLZ_0 := FALSE;
   PouringCycle[1].FLT_Max_Waittime := FALSE;
   PouringCycle[1].FLT_Max_Shottime := FALSE;
   PouringCycle[1].FLT_OP_Mode := FALSE;
   PouringCycle[1].Reserve1 := FALSE;
   PouringCycle[1].Reserve2 := FALSE;
   PouringCycle[1].Reserve3 := FALSE;
   PouringCycle[1].FLT_CompAllocation := FALSE;
   PouringCycle[1].FLT_NewNoTooEarly := FALSE;
   PouringCycle[1].FLT_WRongStationNumber := FALSE;
   PouringCycle[1].FLT_WrongToolNumber := FALSE;
   PouringCycle[1].FLT_WrongShotNumber := FALSE;
   PouringCycle[1].FLT_WrongMixingheadNumber := FALSE;
   PouringCycle[1].FLT_TransferShotResult := FALSE;
   PouringCycle[1].FLT_BufferShotResultFull := FALSE;
   PouringCycle[1].Spare_1_7 := FALSE;
   PouringCycle[2].FLT_KLZ_0 := FALSE;
   PouringCycle[2].FLT_Max_Waittime := FALSE;
   PouringCycle[2].FLT_Max_Shottime := FALSE;
   PouringCycle[2].FLT_OP_Mode := FALSE;
   PouringCycle[2].Reserve1 := FALSE;
   PouringCycle[2].Reserve2 := FALSE;
   PouringCycle[2].Reserve3 := FALSE;
   PouringCycle[2].FLT_CompAllocation := FALSE;
   PouringCycle[2].FLT_NewNoTooEarly := FALSE;
   PouringCycle[2].FLT_WRongStationNumber := FALSE;
   PouringCycle[2].FLT_WrongToolNumber := FALSE;
   PouringCycle[2].FLT_WrongShotNumber := FALSE;
   PouringCycle[2].FLT_WrongMixingheadNumber := FALSE;
   PouringCycle[2].FLT_TransferShotResult := FALSE;
   PouringCycle[2].FLT_BufferShotResultFull := FALSE;
   PouringCycle[2].Spare_1_7 := FALSE;
   Foaming_Time[1].Sensor_FLT_broken_wire := FALSE;
   Foaming_Time[1].Warning_limit_plus := FALSE;
   Foaming_Time[1].Warning_limit_minus := FALSE;
   Foaming_Time[1].Alarm_limit_plus := FALSE;
   Foaming_Time[1].Alarm_limit_minus := FALSE;
   Foaming_Time[1].Controller_at_limit := FALSE;
   Foaming_Time[1].Spare_0_6 := FALSE;
   Foaming_Time[1].Fuse_TemperingOverLoad := FALSE;
   Foaming_Time[1].Spare_1_0 := FALSE;
   Foaming_Time[1].Spare_1_1 := FALSE;
   Foaming_Time[1].Spare_1_2 := FALSE;
   Foaming_Time[1].Spare_1_3 := FALSE;
   Foaming_Time[1].Spare_1_4 := FALSE;
   Foaming_Time[1].Spare_1_5 := FALSE;
   Foaming_Time[1].Spare_1_6 := FALSE;
   Foaming_Time[1].Spare_1_7 := FALSE;
   Foaming_Time[2].Sensor_FLT_broken_wire := FALSE;
   Foaming_Time[2].Warning_limit_plus := FALSE;
   Foaming_Time[2].Warning_limit_minus := FALSE;
   Foaming_Time[2].Alarm_limit_plus := FALSE;
   Foaming_Time[2].Alarm_limit_minus := FALSE;
   Foaming_Time[2].Controller_at_limit := FALSE;
   Foaming_Time[2].Spare_0_6 := FALSE;
   Foaming_Time[2].Fuse_TemperingOverLoad := FALSE;
   Foaming_Time[2].Spare_1_0 := FALSE;
   Foaming_Time[2].Spare_1_1 := FALSE;
   Foaming_Time[2].Spare_1_2 := FALSE;
   Foaming_Time[2].Spare_1_3 := FALSE;
   Foaming_Time[2].Spare_1_4 := FALSE;
   Foaming_Time[2].Spare_1_5 := FALSE;
   Foaming_Time[2].Spare_1_6 := FALSE;
   Foaming_Time[2].Spare_1_7 := FALSE;
END_DATA_BLOCK

DATA_BLOCK "DB900_ConfCalibFlow"   // DB900
TITLE = Configuration max flow calculation
{ S7_Optimized_Access := 'FALSE' }
VERSION : 0.1
   VAR
      ReadWriteDeviceNo : Int := 0;
      CopyDeviceNO : Int := 0;
      Read : Bool := FALSE;
      Write : Bool := FALSE;
      Copy : Bool := FALSE;
      Flow : Array[0..16] of "UDT900_ConfCalibFlow";
   END_VAR
BEGIN
   Flow[1].Density := 1055;
   Flow[3].Density := 880;
   Flow[4].Density := 880;
   Flow[7].Density := 880;
   Flow[8].Density := 880;
   Flow[9].Density := 880;
   Flow[11].Density := 880;
   Flow[13].Density := 1050;
   Flow[15].Density := 1050;
   Flow[1].Pulse_per_liter := 333.0;
   Flow[4].Pulse_per_liter := 965.0;
   Flow[7].Pulse_per_liter := 965.0;
   Flow[8].Pulse_per_liter := 965.0;
   Flow[9].Pulse_per_liter := 965.0;
   Flow[11].Pulse_per_liter := 965.0;
   Flow[13].Pulse_per_liter := 0.0;
   Flow[15].Pulse_per_liter := 0.0;
   Flow[1].MaxFlow := 703.3333;
   Flow[4].MaxFlow := 0.0;
   Flow[7].MaxFlow := 26796.0;
   Flow[8].MaxFlow := 26796.0;
   Flow[9].MaxFlow := 26796.0;
   Flow[11].MaxFlow := 26796.0;
   Flow[13].MaxFlow := 0.0;
   Flow[15].MaxFlow := 0.0;
   Flow[0].Density := 0;
   Flow[0].Pulse_per_liter := 0.0;
   Flow[0].MaxFlow := 0.0;
   Flow[2].Density := 1055;
   Flow[2].Pulse_per_liter := 965.0;
   Flow[2].MaxFlow := 281.3333;
   Flow[3].Pulse_per_liter := 965.0;
   Flow[3].MaxFlow := 0.0;
   Flow[5].Density := 880;
   Flow[5].Pulse_per_liter := 965.0;
   Flow[5].MaxFlow := 26796.0;
   Flow[6].Density := 880;
   Flow[6].Pulse_per_liter := 965.0;
   Flow[6].MaxFlow := 26796.0;
   Flow[10].Density := 880;
   Flow[10].Pulse_per_liter := 965.0;
   Flow[10].MaxFlow := 26796.0;
   Flow[12].Density := 880;
   Flow[12].Pulse_per_liter := 965.0;
   Flow[12].MaxFlow := 26796.0;
   Flow[14].Density := 0;
   Flow[14].Pulse_per_liter := 0.0;
   Flow[14].MaxFlow := 0.0;
   Flow[16].Density := 0;
   Flow[16].Pulse_per_liter := 0.0;
   Flow[16].MaxFlow := 0.0;
   Flow[0].Factor := 0.0;
   Flow[1].Factor := 1.0;
   Flow[2].Factor := 1.0;
   Flow[3].Factor := 0.0;
   Flow[4].Factor := 0.0;
   Flow[5].Factor := 0.0;
   Flow[6].Factor := 0.0;
   Flow[7].Factor := 0.0;
   Flow[8].Factor := 0.0;
   Flow[9].Factor := 0.0;
   Flow[10].Factor := 0.0;
   Flow[11].Factor := 0.0;
   Flow[12].Factor := 0.0;
   Flow[13].Factor := 0.0;
   Flow[14].Factor := 0.0;
   Flow[15].Factor := 0.0;
   Flow[16].Factor := 0.0;
END_DATA_BLOCK

DATA_BLOCK "DB902_ConfFlow_PV"   // DB902
TITLE = Configuration flow values -> ProCan
{ S7_Optimized_Access := 'FALSE' }
VERSION : 0.1
   VAR
      ReadWriteDeviceNo : Int := 1;
      CopyDeviceNO : Int := 0;
      Read : Bool := FALSE;
      Write : Bool := FALSE;
      Copy : Bool := FALSE;
      FlowConf : Array[0..16] of Bool;   // Bit selects flow-number and activates transfer of configuration to ProCan
      Flow : Array[0..16] of "UDT902_ConfFlow";
   END_VAR
BEGIN
   Flow[0].calibration := 10152;
   Flow[1].calibration := 10880;
   Flow[2].calibration := 2572;
   Flow[3].calibration := 0;
   Flow[4].calibration := 0;
   Flow[5].calibration := 0;
   Flow[6].calibration := 0;
   Flow[7].calibration := 0;
   Flow[8].calibration := 0;
   Flow[0].maximumflow := 26667;
   Flow[1].maximumflow := 13333;
   Flow[2].maximumflow := 13333;
   Flow[3].maximumflow := 26796;
   Flow[4].maximumflow := 26796;
   Flow[5].maximumflow := 26796;
   Flow[6].maximumflow := 26796;
   Flow[7].maximumflow := 26796;
   Flow[8].maximumflow := 26796;
   Flow[0].controltime := 200;
   Flow[1].controltime := 200;
   Flow[2].controltime := 200;
   Flow[3].controltime := 100;
   Flow[4].controltime := 100;
   Flow[5].controltime := 100;
   Flow[6].controltime := 100;
   Flow[7].controltime := 100;
   Flow[8].controltime := 100;
   Flow[2].controltime_FPB := 200;
   Flow[1].maximumVoltage := 32760;
   Flow[2].maximumVoltage := 32760;
   Flow[1].single_phase := TRUE;
   Flow[2].single_phase := TRUE;
   Flow[1].controltime_FPB := 200;
   FlowConf[0] := FALSE;
   FlowConf[1] := FALSE;
   FlowConf[2] := FALSE;
   FlowConf[3] := FALSE;
   FlowConf[4] := FALSE;
   FlowConf[5] := FALSE;
   FlowConf[6] := FALSE;
   FlowConf[7] := FALSE;
   FlowConf[8] := FALSE;
   FlowConf[9] := FALSE;
   FlowConf[10] := FALSE;
   FlowConf[11] := FALSE;
   FlowConf[12] := FALSE;
   FlowConf[13] := FALSE;
   FlowConf[14] := FALSE;
   FlowConf[15] := FALSE;
   FlowConf[16] := FALSE;
   Flow[0].Spare_2_0 := FALSE;
   Flow[0].Spare_2_1 := FALSE;
   Flow[0].Spare_2_2 := FALSE;
   Flow[0].Spare_2_3 := FALSE;
   Flow[0].Spare_2_4 := FALSE;
   Flow[0].Spare_2_5 := FALSE;
   Flow[0].Spare_2_6 := FALSE;
   Flow[0].Spare_2_7 := FALSE;
   Flow[0].single_phase := TRUE;
   Flow[0].FPB_SPC0 := FALSE;
   Flow[0].FPB_SPC01 := FALSE;
   Flow[0].Pos_OUT := FALSE;
   Flow[0].Spare_3_04 := FALSE;
   Flow[0].Spare_3_05 := FALSE;
   Flow[0].Spare_3_06 := FALSE;
   Flow[0].Spare_3_07 := FALSE;
   Flow[0].controltime_FPB := 200;
   Flow[0].time_average := 200;
   Flow[0].minimumVoltage := 0;
   Flow[0].maximumVoltage := 32760;
   Flow[0].delayWarn_minVoltage := 5000;
   Flow[0].delayWarn_maxVoltage := 5000;
   Flow[1].Spare_2_0 := FALSE;
   Flow[1].Spare_2_1 := FALSE;
   Flow[1].Spare_2_2 := FALSE;
   Flow[1].Spare_2_3 := FALSE;
   Flow[1].Spare_2_4 := FALSE;
   Flow[1].Spare_2_5 := FALSE;
   Flow[1].Spare_2_6 := FALSE;
   Flow[1].Spare_2_7 := FALSE;
   Flow[1].FPB_SPC0 := FALSE;
   Flow[1].FPB_SPC01 := FALSE;
   Flow[1].Pos_OUT := FALSE;
   Flow[1].Spare_3_04 := FALSE;
   Flow[1].Spare_3_05 := FALSE;
   Flow[1].Spare_3_06 := FALSE;
   Flow[1].Spare_3_07 := FALSE;
   Flow[1].time_average := 200;
   Flow[1].minimumVoltage := 0;
   Flow[1].delayWarn_minVoltage := 5000;
   Flow[1].delayWarn_maxVoltage := 5000;
   Flow[2].Spare_2_0 := FALSE;
   Flow[2].Spare_2_1 := FALSE;
   Flow[2].Spare_2_2 := FALSE;
   Flow[2].Spare_2_3 := FALSE;
   Flow[2].Spare_2_4 := FALSE;
   Flow[2].Spare_2_5 := FALSE;
   Flow[2].Spare_2_6 := FALSE;
   Flow[2].Spare_2_7 := FALSE;
   Flow[2].FPB_SPC0 := FALSE;
   Flow[2].FPB_SPC01 := FALSE;
   Flow[2].Pos_OUT := FALSE;
   Flow[2].Spare_3_04 := FALSE;
   Flow[2].Spare_3_05 := FALSE;
   Flow[2].Spare_3_06 := FALSE;
   Flow[2].Spare_3_07 := FALSE;
   Flow[2].time_average := 200;
   Flow[2].minimumVoltage := 0;
   Flow[2].delayWarn_minVoltage := 5000;
   Flow[2].delayWarn_maxVoltage := 5000;
   Flow[3].Spare_2_0 := FALSE;
   Flow[3].Spare_2_1 := FALSE;
   Flow[3].Spare_2_2 := FALSE;
   Flow[3].Spare_2_3 := FALSE;
   Flow[3].Spare_2_4 := FALSE;
   Flow[3].Spare_2_5 := FALSE;
   Flow[3].Spare_2_6 := FALSE;
   Flow[3].Spare_2_7 := FALSE;
   Flow[3].single_phase := FALSE;
   Flow[3].FPB_SPC0 := FALSE;
   Flow[3].FPB_SPC01 := FALSE;
   Flow[3].Pos_OUT := FALSE;
   Flow[3].Spare_3_04 := FALSE;
   Flow[3].Spare_3_05 := FALSE;
   Flow[3].Spare_3_06 := FALSE;
   Flow[3].Spare_3_07 := FALSE;
   Flow[3].controltime_FPB := 500;
   Flow[3].time_average := 200;
   Flow[3].minimumVoltage := 0;
   Flow[3].maximumVoltage := 32767;
   Flow[3].delayWarn_minVoltage := 5000;
   Flow[3].delayWarn_maxVoltage := 5000;
   Flow[4].Spare_2_0 := FALSE;
   Flow[4].Spare_2_1 := FALSE;
   Flow[4].Spare_2_2 := FALSE;
   Flow[4].Spare_2_3 := FALSE;
   Flow[4].Spare_2_4 := FALSE;
   Flow[4].Spare_2_5 := FALSE;
   Flow[4].Spare_2_6 := FALSE;
   Flow[4].Spare_2_7 := FALSE;
   Flow[4].single_phase := FALSE;
   Flow[4].FPB_SPC0 := FALSE;
   Flow[4].FPB_SPC01 := FALSE;
   Flow[4].Pos_OUT := FALSE;
   Flow[4].Spare_3_04 := FALSE;
   Flow[4].Spare_3_05 := FALSE;
   Flow[4].Spare_3_06 := FALSE;
   Flow[4].Spare_3_07 := FALSE;
   Flow[4].controltime_FPB := 500;
   Flow[4].time_average := 200;
   Flow[4].minimumVoltage := 0;
   Flow[4].maximumVoltage := 32767;
   Flow[4].delayWarn_minVoltage := 5000;
   Flow[4].delayWarn_maxVoltage := 5000;
   Flow[5].Spare_2_0 := FALSE;
   Flow[5].Spare_2_1 := FALSE;
   Flow[5].Spare_2_2 := FALSE;
   Flow[5].Spare_2_3 := FALSE;
   Flow[5].Spare_2_4 := FALSE;
   Flow[5].Spare_2_5 := FALSE;
   Flow[5].Spare_2_6 := FALSE;
   Flow[5].Spare_2_7 := FALSE;
   Flow[5].single_phase := FALSE;
   Flow[5].FPB_SPC0 := FALSE;
   Flow[5].FPB_SPC01 := FALSE;
   Flow[5].Pos_OUT := FALSE;
   Flow[5].Spare_3_04 := FALSE;
   Flow[5].Spare_3_05 := FALSE;
   Flow[5].Spare_3_06 := FALSE;
   Flow[5].Spare_3_07 := FALSE;
   Flow[5].controltime_FPB := 500;
   Flow[5].time_average := 200;
   Flow[5].minimumVoltage := 0;
   Flow[5].maximumVoltage := 32767;
   Flow[5].delayWarn_minVoltage := 5000;
   Flow[5].delayWarn_maxVoltage := 5000;
   Flow[6].Spare_2_0 := FALSE;
   Flow[6].Spare_2_1 := FALSE;
   Flow[6].Spare_2_2 := FALSE;
   Flow[6].Spare_2_3 := FALSE;
   Flow[6].Spare_2_4 := FALSE;
   Flow[6].Spare_2_5 := FALSE;
   Flow[6].Spare_2_6 := FALSE;
   Flow[6].Spare_2_7 := FALSE;
   Flow[6].single_phase := FALSE;
   Flow[6].FPB_SPC0 := FALSE;
   Flow[6].FPB_SPC01 := FALSE;
   Flow[6].Pos_OUT := FALSE;
   Flow[6].Spare_3_04 := FALSE;
   Flow[6].Spare_3_05 := FALSE;
   Flow[6].Spare_3_06 := FALSE;
   Flow[6].Spare_3_07 := FALSE;
   Flow[6].controltime_FPB := 500;
   Flow[6].time_average := 200;
   Flow[6].minimumVoltage := 0;
   Flow[6].maximumVoltage := 32767;
   Flow[6].delayWarn_minVoltage := 5000;
   Flow[6].delayWarn_maxVoltage := 5000;
   Flow[7].Spare_2_0 := FALSE;
   Flow[7].Spare_2_1 := FALSE;
   // 242 more start values not shown
END_DATA_BLOCK

DATA_BLOCK "DB917_ShotResult5"   // DB917
{ S7_Optimized_Access := 'TRUE' }
VERSION : 0.1
   VAR RETAIN
      Start : Int;
      StartDate : Date;
      StartTime : Time_Of_Day;
      Shots : Array[1..5] of "UDT927_ShotResult5";
   END_VAR
BEGIN
END_DATA_BLOCK

DATA_BLOCK "DB918_ShotResultlast10"   // DB918
{ S7_Optimized_Access := 'FALSE' }